REGION Network 13: Manual mode request
   RUNG wire#powerrail
      Contact( "Z256".ST_xSelectionManualMode )
      I_Contact( "Z256".ST_xManualModeAccepted )
      Coil( "Z256".ST_xManualModeRequest )
   END_RUNG
   // the same network as SCL:
   "Z256".ST_xManualModeRequest := "Z256".ST_xSelectionManualMode AND NOT "Z256".ST_xManualModeAccepted;
END_REGION

REGION Network 14: Manual mode accepted
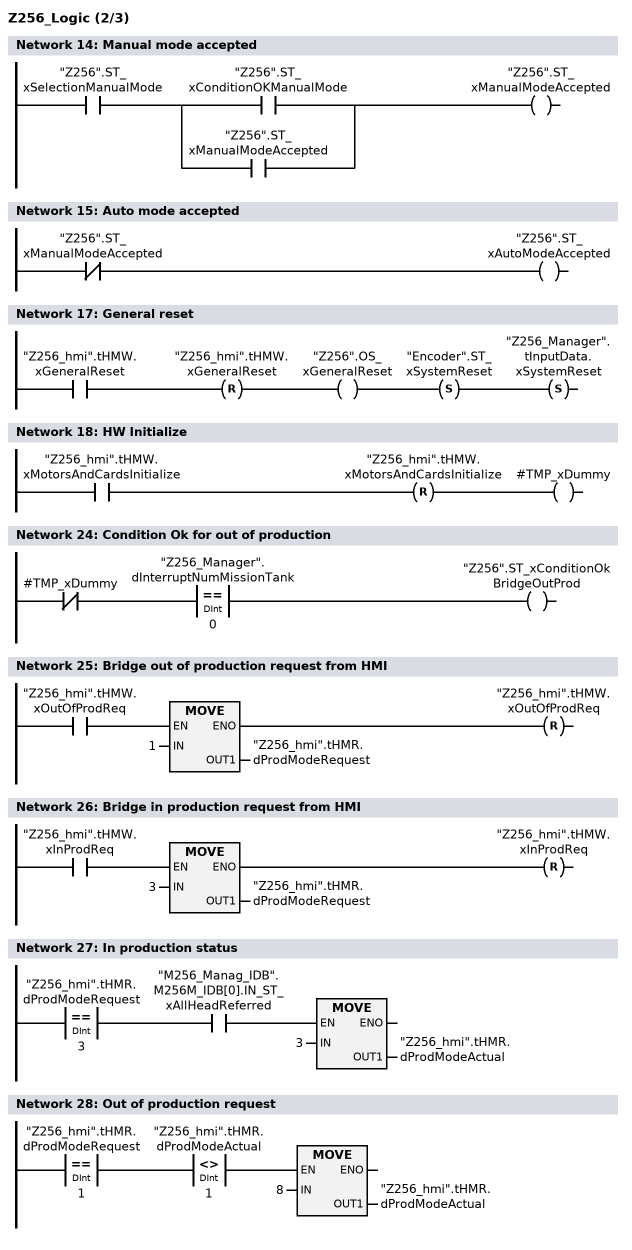
   RUNG wire#powerrail
      Contact( "Z256".ST_xSelectionManualMode )
      wire#w1
      Contact( "Z256".ST_xConditionOKManualMode )
      wire#w2
      Coil( "Z256".ST_xManualModeAccepted )
   END_RUNG
   RUNG wire#w1
      Contact( "Z256".ST_xManualModeAccepted )
   END_RUNG wire#w2
   // the same network as SCL:
   "Z256".ST_xManualModeAccepted := "Z256".ST_xSelectionManualMode AND ("Z256".ST_xConditionOKManualMode OR "Z256".ST_xManualModeAccepted);
END_REGION

REGION Network 15: Auto mode accepted
   RUNG wire#powerrail
      I_Contact( "Z256".ST_xManualModeAccepted )
      Coil( "Z256".ST_xAutoModeAccepted )
   END_RUNG
   // the same network as SCL:
   "Z256".ST_xAutoModeAccepted := NOT "Z256".ST_xManualModeAccepted;
END_REGION

REGION Network 16: ### HMI LOGICS ###
END_REGION

REGION Network 17: General reset
   RUNG wire#powerrail
      Contact( "Z256_hmi".tHMW.xGeneralReset )
      R_Coil( "Z256_hmi".tHMW.xGeneralReset )
      Coil( "Z256".OS_xGeneralReset )
      S_Coil( "Encoder".ST_xSystemReset )
      S_Coil( "Z256_Manager".tInputData.xSystemReset )
   END_RUNG
   // the same network as SCL:
   #_w1 := "Z256_hmi".tHMW.xGeneralReset;
   IF #_w1 THEN "Z256_hmi".tHMW.xGeneralReset := FALSE; END_IF;
   "Z256".OS_xGeneralReset := #_w1;
   IF #_w1 THEN
       "Encoder".ST_xSystemReset := TRUE;
       "Z256_Manager".tInputData.xSystemReset := TRUE;
   END_IF;
END_REGION

REGION Network 18: HW Initialize
   RUNG wire#powerrail
      Contact( "Z256_hmi".tHMW.xMotorsAndCardsInitialize )
      R_Coil( "Z256_hmi".tHMW.xMotorsAndCardsInitialize )
      Coil( #TMP_xDummy )
   END_RUNG
   // the same network as SCL:
   #_w1 := "Z256_hmi".tHMW.xMotorsAndCardsInitialize;
   IF #_w1 THEN "Z256_hmi".tHMW.xMotorsAndCardsInitialize := FALSE; END_IF;
   #TMP_xDummy := #_w1;
END_REGION

REGION Network 19 (SCL): Reset head initialized
   IF #TMP_xDummy THEN

       FOR #TMP_iIndex := 0 TO "CONST_dNumberOfHeadsCycle" BY 1
       DO
           "M256_Manag_IDB".M256M_IDB[#TMP_iIndex].ST_xHeadInitialized := 0;
       END_FOR;

   END_IF;
END_REGION

REGION Network 20: Cut with glass break
   // tolto enable /disable , messo che scada lo mette ad ON/OFF
END_REGION

REGION Network 21 (SCL): Enable/disable head from scada
    //   FOR #TMP_iIndex := 0 TO "CONST_dNumberOfHeadsCycle" DO
    //       IF "Z256_hmi".tHMW.rgxEnableHead[#TMP_iIndex] THEN
     //          "Z256_hmi".tHMW.rgxEnableHead[#TMP_iIndex] := 0;
     //          "Z256_hmi".tHMR.rgxHeadEnabled[#TMP_iIndex] := 1;
    //       END_IF;
    //       IF "Z256_hmi".tHMW.rgxDisableHead[#TMP_iIndex] THEN
    //           "Z256_hmi".tHMW.rgxDisableHead[#TMP_iIndex] := 0;
    //           "Z256_hmi".tHMR.rgxHeadEnabled[#TMP_iIndex] := 0;
    //       END_IF;
    //   END_FOR;
END_REGION

REGION Network 22: ### PRODUCTIONS STATUS ###
END_REGION

REGION Network 23 (SCL)
   #TMP_xDummy := false;
   FOR #TMP_iIndex:=0 TO "CONST_dNumberOfHeadsCycle" DO
       IF "Z256_Manager".tOutputData.rgxDataToProcessInter[#TMP_iIndex]=TRUE THEN
           #TMP_xDummy := true;
       END_IF;
   END_FOR;
END_REGION

REGION Network 24: Condition Ok for out of production
   RUNG wire#powerrail
      I_Contact( #TMP_xDummy )
      { S7_Templates := "SrcType := DInt" } EQ_Contact(in1 := "Z256_Manager".dInterruptNumMissionTank, in2 := 0)
      Coil( "Z256".ST_xConditionOkBridgeOutProd )
   END_RUNG
   // the same network as SCL:
   "Z256".ST_xConditionOkBridgeOutProd := NOT #TMP_xDummy AND ("Z256_Manager".dInterruptNumMissionTank = 0);
END_REGION

REGION Network 25: Bridge out of production request from HMI
   RUNG wire#powerrail
      Contact( "Z256_hmi".tHMW.xOutOfProdReq )
      Move(in := 1, out1 => "Z256_hmi".tHMR.dProdModeRequest)
      R_Coil( "Z256_hmi".tHMW.xOutOfProdReq )
   END_RUNG
   // the same network as SCL:
   IF "Z256_hmi".tHMW.xOutOfProdReq THEN
       "Z256_hmi".tHMR.dProdModeRequest := 1;
       "Z256_hmi".tHMW.xOutOfProdReq := FALSE;
   END_IF;
END_REGION

REGION Network 26: Bridge in production request from HMI
   RUNG wire#powerrail
      Contact( "Z256_hmi".tHMW.xInProdReq )
      Move(in := 3, out1 => "Z256_hmi".tHMR.dProdModeRequest)
      R_Coil( "Z256_hmi".tHMW.xInProdReq )
   END_RUNG
   // the same network as SCL:
   IF "Z256_hmi".tHMW.xInProdReq THEN
       "Z256_hmi".tHMR.dProdModeRequest := 3;
       "Z256_hmi".tHMW.xInProdReq := FALSE;
   END_IF;
END_REGION

REGION Network 27: In production status
   RUNG wire#powerrail
      { S7_Templates := "SrcType := DInt" } EQ_Contact(in1 := "Z256_hmi".tHMR.dProdModeRequest, in2 := 3)
      Contact( "M256_Manag_IDB".M256M_IDB[0].IN_ST_xAllHeadReferred )
      Move(in := 3, out1 => "Z256_hmi".tHMR.dProdModeActual)
   END_RUNG
   // the same network as SCL:
   IF ("Z256_hmi".tHMR.dProdModeRequest = 3) AND "M256_Manag_IDB".M256M_IDB[0].IN_ST_xAllHeadReferred THEN
       "Z256_hmi".tHMR.dProdModeActual := 3;
   END_IF;
END_REGION

REGION Network 28: Out of production request
   RUNG wire#powerrail
      { S7_Templates := "SrcType := DInt" } EQ_Contact(in1 := "Z256_hmi".tHMR.dProdModeRequest, in2 := 1)
      { S7_Templates := "SrcType := DInt" } NE_Contact(in1 := "Z256_hmi".tHMR.dProdModeActual, in2 := 1)
      Move(in := 8, out1 => "Z256_hmi".tHMR.dProdModeActual)
   END_RUNG
   // the same network as SCL:
   IF ("Z256_hmi".tHMR.dProdModeRequest = 1) AND ("Z256_hmi".tHMR.dProdModeActual <> 1) THEN
       "Z256_hmi".tHMR.dProdModeActual := 8;
   END_IF;
END_REGION

REGION Network 29: Out of production status
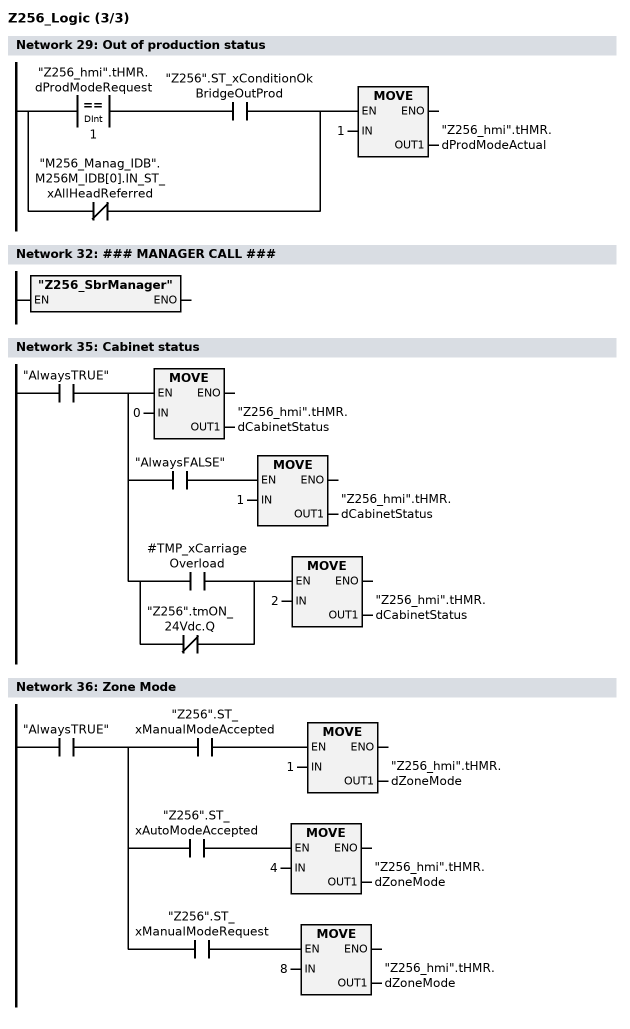
   RUNG wire#powerrail
      { S7_Templates := "SrcType := DInt" } EQ_Contact(in1 := "Z256_hmi".tHMR.dProdModeRequest, in2 := 1)
      Contact( "Z256".ST_xConditionOkBridgeOutProd )
      wire#w1
      Move(in := 1, out1 => "Z256_hmi".tHMR.dProdModeActual)
   END_RUNG
   RUNG wire#powerrail
      I_Contact( "M256_Manag_IDB".M256M_IDB[0].IN_ST_xAllHeadReferred )
   END_RUNG wire#w1
   // the same network as SCL:
   IF (("Z256_hmi".tHMR.dProdModeRequest = 1) AND "Z256".ST_xConditionOkBridgeOutProd) OR NOT "M256_Manag_IDB".M256M_IDB[0].IN_ST_xAllHeadReferred THEN
       "Z256_hmi".tHMR.dProdModeActual := 1;
   END_IF;
END_REGION

REGION Network 30 (SCL): Calculate head status

   FOR #TMP_iIndex := 0 TO "CONST_dNumberOfHeadsCycle" BY 1
   DO
       "Z256_SbrHeadsStatuses"(#TMP_iIndex);
   END_FOR;
END_REGION

REGION Network 31 (SCL): Reset head referred after emergency
   FOR #TMP_iIndex := 0 TO "CONST_dNumberOfHeadsCycle" DO
       IF "DB_Z256_Scada".tAlm.tE.x0 OR "DB_Z256_Scada".tAlm.tE.x1 OR NOT("M256_Manag_IDB".M256M_IDB[#TMP_iIndex].INPUT_xCarriageOverload) THEN
           "M256_Manag_IDB".M256M_IDB[#TMP_iIndex].ST_xHeadReferredSwitch := 0;
       END_IF;
   END_FOR;
END_REGION

REGION Network 32: ### MANAGER CALL ###
   RUNG wire#powerrail
      "Z256_SbrManager"()
   END_RUNG
   // the same network as SCL:
   "Z256_SbrManager"();
END_REGION

REGION Network 33: #### HMI STATUS ####
END_REGION

REGION Network 34 (SCL): Carriage overload array check
   #TMP_xCarriageOverload := false;
   FOR #TMP_iIndex := 0 TO "CONST_dNumberOfHeadsCycle" DO
       IF "M256_Manag_IDB".M256M_IDB[#TMP_iIndex].tALM.tS.x3 THEN
           #TMP_xCarriageOverload := true;
       END_IF;
   END_FOR;
END_REGION

REGION Network 35: Cabinet status
   RUNG wire#powerrail
      Contact( "AlwaysTRUE" )
      wire#w1
      Move(in := 0, out1 => "Z256_hmi".tHMR.dCabinetStatus)
   END_RUNG
   RUNG wire#w1
      Contact( "AlwaysFALSE" )
      Move(in := 1, out1 => "Z256_hmi".tHMR.dCabinetStatus)
   END_RUNG
   RUNG wire#w1
      Contact( #TMP_xCarriageOverload )
      wire#w2
      Move(in := 2, out1 => "Z256_hmi".tHMR.dCabinetStatus)
   END_RUNG
   RUNG wire#w1
      I_Contact( "Z256".tmON_24Vdc.Q )
   END_RUNG wire#w2
   // the same network as SCL:
   IF "AlwaysTRUE" THEN "Z256_hmi".tHMR.dCabinetStatus := 0; END_IF;
   IF "AlwaysTRUE" AND "AlwaysFALSE" THEN "Z256_hmi".tHMR.dCabinetStatus := 1; END_IF;
   IF "AlwaysTRUE" AND (#TMP_xCarriageOverload OR NOT "Z256".tmON_24Vdc.Q) THEN
       "Z256_hmi".tHMR.dCabinetStatus := 2;
   END_IF;
END_REGION

REGION Network 36: Zone Mode
   RUNG wire#powerrail
      Contact( "AlwaysTRUE" )
      wire#w1
      Contact( "Z256".ST_xManualModeAccepted )
      Move(in := 1, out1 => "Z256_hmi".tHMR.dZoneMode)
   END_RUNG
   RUNG wire#w1
      Contact( "Z256".ST_xAutoModeAccepted )
      Move(in := 4, out1 => "Z256_hmi".tHMR.dZoneMode)
   END_RUNG
   RUNG wire#w1
      Contact( "Z256".ST_xManualModeRequest )
      Move(in := 8, out1 => "Z256_hmi".tHMR.dZoneMode)
   END_RUNG
   // the same network as SCL:
   IF "AlwaysTRUE" AND "Z256".ST_xManualModeAccepted THEN "Z256_hmi".tHMR.dZoneMode := 1; END_IF;
   IF "AlwaysTRUE" AND "Z256".ST_xAutoModeAccepted THEN "Z256_hmi".tHMR.dZoneMode := 4; END_IF;
   IF "AlwaysTRUE" AND "Z256".ST_xManualModeRequest THEN "Z256_hmi".tHMR.dZoneMode := 8; END_IF;
END_REGION

REGION Network 37 (SCL): Set all brake engage/release
   IF "Z256_hmi".tHMW.tManCmd.xBrakeEngage THEN
       FOR #TMP_iIndex := 0 TO "CONST_dNumberOfHeadsCycle" BY 1
       DO
           "M256_Manag_IDB".M256M_IDB[#TMP_iIndex].tHMW.xBrakeEngageHeads := 1;
       END_FOR;
       "Z256_hmi".tHMW.tManCmd.xBrakeEngage := 0;
   END_IF;
   IF "Z256_hmi".tHMW.tManCmd.xBrakeRelease THEN
       FOR #TMP_iIndex := 0 TO "CONST_dNumberOfHeadsCycle" BY 1
       DO
           "M256_Manag_IDB".M256M_IDB[#TMP_iIndex].tHMW.xBrakeRealeaseHeads := 1;
       END_FOR;
       "Z256_hmi".tHMW.tManCmd.xBrakeRelease := 0;
   END_IF;
END_REGION
END_FUNCTION

FUNCTION "Z256_Faults" : Void   // FC3, LAD
{ S7_Optimized_Access := 'TRUE' }
VERSION : 0.1
   VAR_TEMP
      TMP_dIndex : DInt;
      TMP_dwDummy : DWord;
      TMP_dwDummy_1 : DWord;
      TMP_dwDummy_2 : DWord;
      TMP_dwDummy_3 : DWord;
      TMP_idummy : Int;
   END_VAR
   VAR_TEMP   // added for the SCL form of the ladder/FBD networks
      _w1 : Bool;
   END_VAR
BEGIN

REGION Network 1: ##### FAULTS #####
END_REGION

REGION Network 2: Reset faults
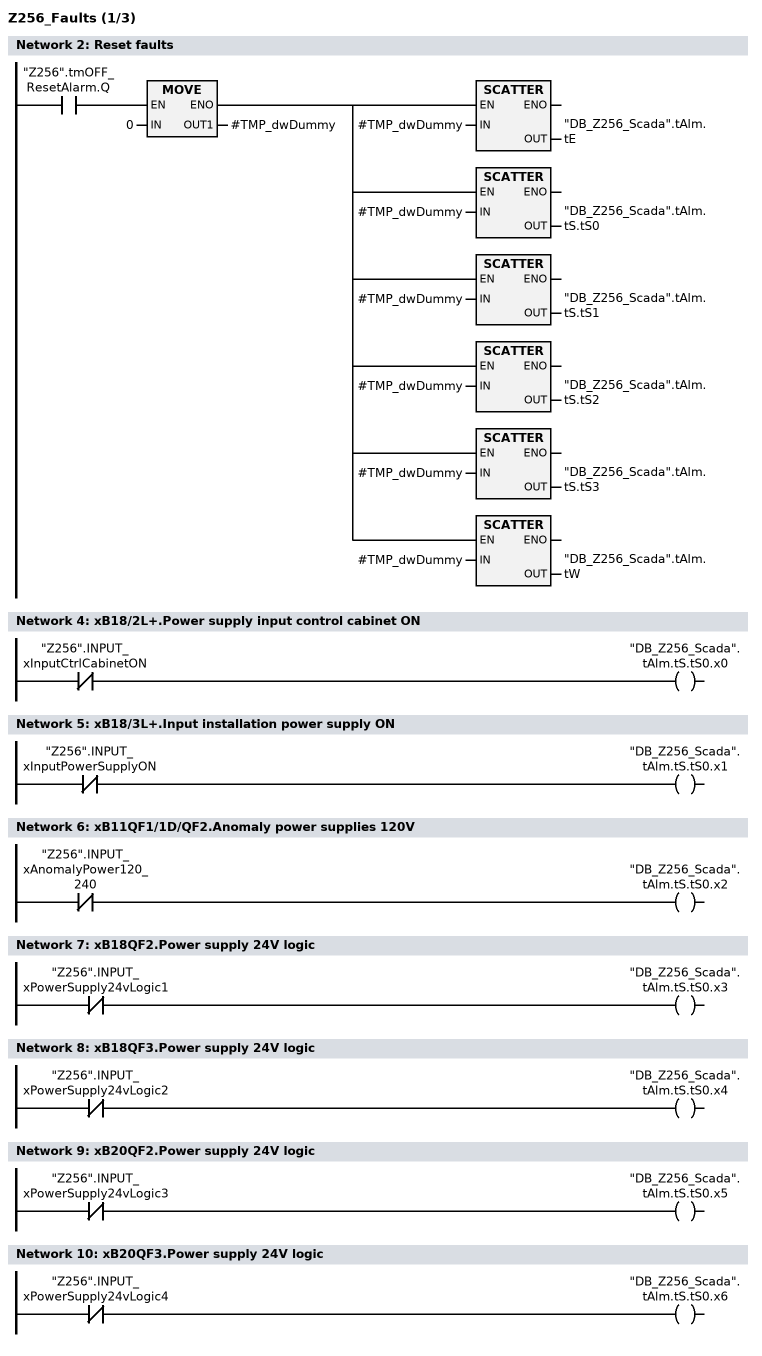
   IF "Z256".tmOFF_ResetAlarm.Q THEN #TMP_dwDummy := 0; END_IF;
   #_w1 := "Z256".tmOFF_ResetAlarm.Q;
   IF #_w1 THEN
       SCATTER(IN := #TMP_dwDummy, OUT => "DB_Z256_Scada".tAlm.tE);
       SCATTER(IN := #TMP_dwDummy, OUT => "DB_Z256_Scada".tAlm.tS.tS0);
       SCATTER(IN := #TMP_dwDummy, OUT => "DB_Z256_Scada".tAlm.tS.tS1);
       SCATTER(IN := #TMP_dwDummy, OUT => "DB_Z256_Scada".tAlm.tS.tS2);
       SCATTER(IN := #TMP_dwDummy, OUT => "DB_Z256_Scada".tAlm.tS.tS3);
       SCATTER(IN := #TMP_dwDummy, OUT => "DB_Z256_Scada".tAlm.tW);
   END_IF;
END_REGION

REGION Network 3: ### CABINET POWER FAULTS ###
END_REGION

REGION Network 4: xB18/2L+.Power supply input control cabinet ON
   RUNG wire#powerrail
      I_Contact( "Z256".INPUT_xInputCtrlCabinetON )
      Coil( "DB_Z256_Scada".tAlm.tS.tS0.x0 )
   END_RUNG
   // the same network as SCL:
   "DB_Z256_Scada".tAlm.tS.tS0.x0 := NOT "Z256".INPUT_xInputCtrlCabinetON;
END_REGION

REGION Network 5: xB18/3L+.Input installation power supply ON
   RUNG wire#powerrail
      I_Contact( "Z256".INPUT_xInputPowerSupplyON )
      Coil( "DB_Z256_Scada".tAlm.tS.tS0.x1 )
   END_RUNG
   // the same network as SCL:
   "DB_Z256_Scada".tAlm.tS.tS0.x1 := NOT "Z256".INPUT_xInputPowerSupplyON;
END_REGION

REGION Network 6: xB11QF1/1D/QF2.Anomaly power supplies 120V
   RUNG wire#powerrail
      I_Contact( "Z256".INPUT_xAnomalyPower120_240 )
      Coil( "DB_Z256_Scada".tAlm.tS.tS0.x2 )
   END_RUNG
   // the same network as SCL:
   "DB_Z256_Scada".tAlm.tS.tS0.x2 := NOT "Z256".INPUT_xAnomalyPower120_240;
END_REGION

REGION Network 7: xB18QF2.Power supply 24V logic
   RUNG wire#powerrail
      I_Contact( "Z256".INPUT_xPowerSupply24vLogic1 )
      Coil( "DB_Z256_Scada".tAlm.tS.tS0.x3 )
   END_RUNG
   // the same network as SCL:
   "DB_Z256_Scada".tAlm.tS.tS0.x3 := NOT "Z256".INPUT_xPowerSupply24vLogic1;
END_REGION

REGION Network 8: xB18QF3.Power supply 24V logic
   RUNG wire#powerrail
      I_Contact( "Z256".INPUT_xPowerSupply24vLogic2 )
      Coil( "DB_Z256_Scada".tAlm.tS.tS0.x4 )
   END_RUNG
   // the same network as SCL:
   "DB_Z256_Scada".tAlm.tS.tS0.x4 := NOT "Z256".INPUT_xPowerSupply24vLogic2;
END_REGION

REGION Network 9: xB20QF2.Power supply 24V logic
   RUNG wire#powerrail
      I_Contact( "Z256".INPUT_xPowerSupply24vLogic3 )
      Coil( "DB_Z256_Scada".tAlm.tS.tS0.x5 )
   END_RUNG
   // the same network as SCL:
   "DB_Z256_Scada".tAlm.tS.tS0.x5 := NOT "Z256".INPUT_xPowerSupply24vLogic3;
END_REGION

REGION Network 10: xB20QF3.Power supply 24V logic
   RUNG wire#powerrail
      I_Contact( "Z256".INPUT_xPowerSupply24vLogic4 )
      Coil( "DB_Z256_Scada".tAlm.tS.tS0.x6 )
   END_RUNG
   // the same network as SCL:
   "DB_Z256_Scada".tAlm.tS.tS0.x6 := NOT "Z256".INPUT_xPowerSupply24vLogic4;
END_REGION

REGION Network 11: xB21QF1.Power supply 24V logic
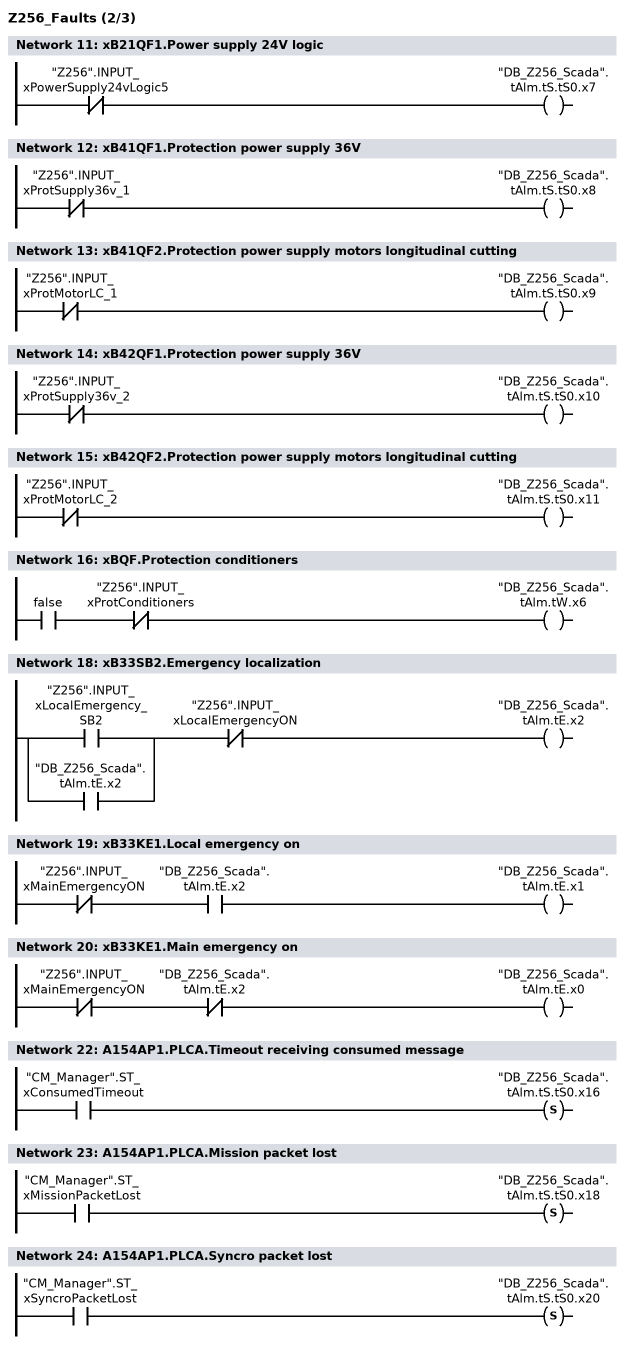
   RUNG wire#powerrail
      I_Contact( "Z256".INPUT_xPowerSupply24vLogic5 )
      Coil( "DB_Z256_Scada".tAlm.tS.tS0.x7 )
   END_RUNG
   // the same network as SCL:
   "DB_Z256_Scada".tAlm.tS.tS0.x7 := NOT "Z256".INPUT_xPowerSupply24vLogic5;
END_REGION

REGION Network 12: xB41QF1.Protection power supply 36V
   RUNG wire#powerrail
      I_Contact( "Z256".INPUT_xProtSupply36v_1 )
      Coil( "DB_Z256_Scada".tAlm.tS.tS0.x8 )
   END_RUNG
   // the same network as SCL:
   "DB_Z256_Scada".tAlm.tS.tS0.x8 := NOT "Z256".INPUT_xProtSupply36v_1;
END_REGION

REGION Network 13: xB41QF2.Protection power supply motors longitudinal cutting
   RUNG wire#powerrail
      I_Contact( "Z256".INPUT_xProtMotorLC_1 )
      Coil( "DB_Z256_Scada".tAlm.tS.tS0.x9 )
   END_RUNG
   // the same network as SCL:
   "DB_Z256_Scada".tAlm.tS.tS0.x9 := NOT "Z256".INPUT_xProtMotorLC_1;
END_REGION

REGION Network 14: xB42QF1.Protection power supply 36V
   RUNG wire#powerrail
      I_Contact( "Z256".INPUT_xProtSupply36v_2 )
      Coil( "DB_Z256_Scada".tAlm.tS.tS0.x10 )
   END_RUNG
   // the same network as SCL:
   "DB_Z256_Scada".tAlm.tS.tS0.x10 := NOT "Z256".INPUT_xProtSupply36v_2;
END_REGION

REGION Network 15: xB42QF2.Protection power supply motors longitudinal cutting
   RUNG wire#powerrail
      I_Contact( "Z256".INPUT_xProtMotorLC_2 )
      Coil( "DB_Z256_Scada".tAlm.tS.tS0.x11 )
   END_RUNG
   // the same network as SCL:
   "DB_Z256_Scada".tAlm.tS.tS0.x11 := NOT "Z256".INPUT_xProtMotorLC_2;
END_REGION

REGION Network 16: xBQF.Protection conditioners
   RUNG wire#powerrail
      Contact( false )
      I_Contact( "Z256".INPUT_xProtConditioners )
      Coil( "DB_Z256_Scada".tAlm.tW.x6 )
   END_RUNG
   // the same network as SCL:
   "DB_Z256_Scada".tAlm.tW.x6 := false AND NOT "Z256".INPUT_xProtConditioners;
END_REGION

REGION Network 17: ### EMERGENCY ###
END_REGION

REGION Network 18: xB33SB2.Emergency localization
   RUNG wire#powerrail
      Contact( "Z256".INPUT_xLocalEmergency_SB2 )
      wire#w1
      I_Contact( "Z256".INPUT_xLocalEmergencyON )
      Coil( "DB_Z256_Scada".tAlm.tE.x2 )
   END_RUNG
   RUNG wire#powerrail
      Contact( "DB_Z256_Scada".tAlm.tE.x2 )
   END_RUNG wire#w1
   // the same network as SCL:
   "DB_Z256_Scada".tAlm.tE.x2 := ("Z256".INPUT_xLocalEmergency_SB2 OR "DB_Z256_Scada".tAlm.tE.x2) AND NOT "Z256".INPUT_xLocalEmergencyON;
END_REGION

REGION Network 19: xB33KE1.Local emergency on
   RUNG wire#powerrail
      I_Contact( "Z256".INPUT_xMainEmergencyON )
      Contact( "DB_Z256_Scada".tAlm.tE.x2 )
      Coil( "DB_Z256_Scada".tAlm.tE.x1 )
   END_RUNG
   // the same network as SCL:
   "DB_Z256_Scada".tAlm.tE.x1 := NOT "Z256".INPUT_xMainEmergencyON AND "DB_Z256_Scada".tAlm.tE.x2;
END_REGION

REGION Network 20: xB33KE1.Main emergency on
   RUNG wire#powerrail
      I_Contact( "Z256".INPUT_xMainEmergencyON )
      I_Contact( "DB_Z256_Scada".tAlm.tE.x2 )
      Coil( "DB_Z256_Scada".tAlm.tE.x0 )
   END_RUNG
   // the same network as SCL:
   "DB_Z256_Scada".tAlm.tE.x0 := NOT "Z256".INPUT_xMainEmergencyON AND NOT "DB_Z256_Scada".tAlm.tE.x2;
END_REGION

REGION Network 21: ### COMMUNICATIONS STOPPING ###
END_REGION

REGION Network 22: A154AP1.PLCA.Timeout receiving consumed message
   RUNG wire#powerrail
      Contact( "CM_Manager".ST_xConsumedTimeout )
      S_Coil( "DB_Z256_Scada".tAlm.tS.tS0.x16 )
   END_RUNG
   // the same network as SCL:
   IF "CM_Manager".ST_xConsumedTimeout THEN "DB_Z256_Scada".tAlm.tS.tS0.x16 := TRUE; END_IF;
END_REGION

REGION Network 23: A154AP1.PLCA.Mission packet lost
   RUNG wire#powerrail
      Contact( "CM_Manager".ST_xMissionPacketLost )
      S_Coil( "DB_Z256_Scada".tAlm.tS.tS0.x18 )
   END_RUNG
   // the same network as SCL:
   IF "CM_Manager".ST_xMissionPacketLost THEN "DB_Z256_Scada".tAlm.tS.tS0.x18 := TRUE; END_IF;
END_REGION

REGION Network 24: A154AP1.PLCA.Syncro packet lost
   RUNG wire#powerrail
      Contact( "CM_Manager".ST_xSyncroPacketLost )
      S_Coil( "DB_Z256_Scada".tAlm.tS.tS0.x20 )
   END_RUNG
   // the same network as SCL:
   IF "CM_Manager".ST_xSyncroPacketLost THEN "DB_Z256_Scada".tAlm.tS.tS0.x20 := TRUE; END_IF;
END_REGION

REGION Network 25: ### SYNCRONIZATION ###
END_REGION

REGION Network 26: Syncro.YCut meter gap outside the limits
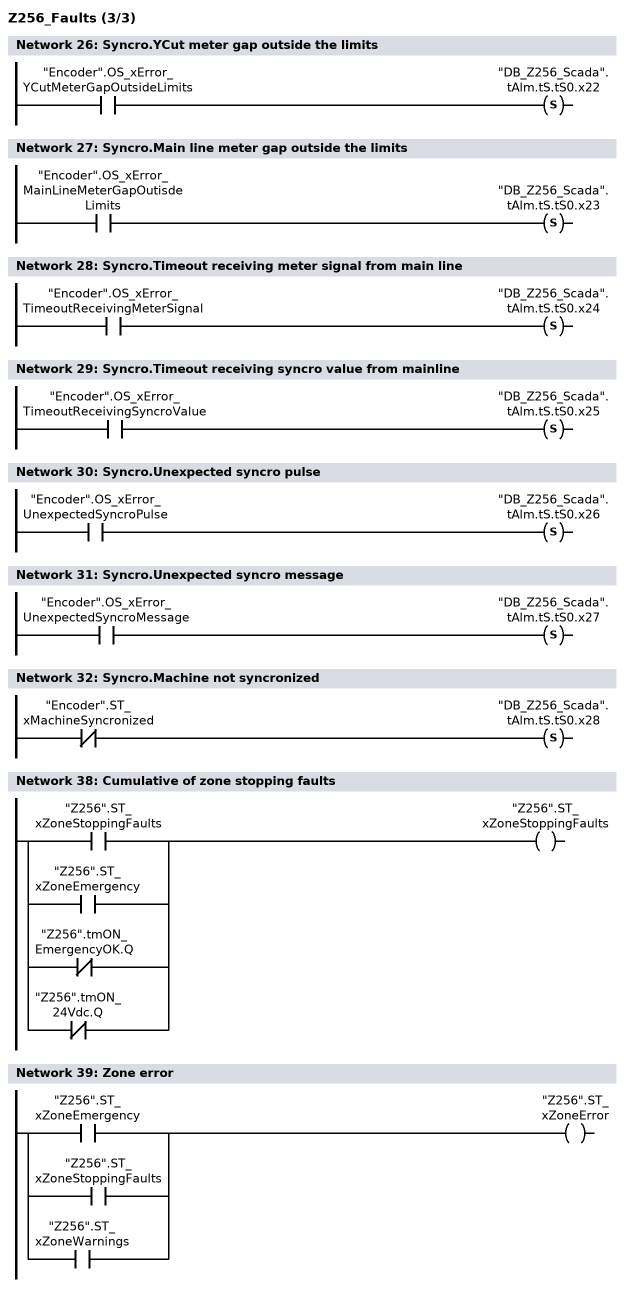
   RUNG wire#powerrail
      Contact( "Encoder".OS_xError_YCutMeterGapOutsideLimits )
      S_Coil( "DB_Z256_Scada".tAlm.tS.tS0.x22 )
   END_RUNG
   // the same network as SCL:
   IF "Encoder".OS_xError_YCutMeterGapOutsideLimits THEN "DB_Z256_Scada".tAlm.tS.tS0.x22 := TRUE; END_IF;
END_REGION

REGION Network 27: Syncro.Main line meter gap outside the limits
   RUNG wire#powerrail
      Contact( "Encoder".OS_xError_MainLineMeterGapOutisdeLimits )
      S_Coil( "DB_Z256_Scada".tAlm.tS.tS0.x23 )
   END_RUNG
   // the same network as SCL:
   IF "Encoder".OS_xError_MainLineMeterGapOutisdeLimits THEN "DB_Z256_Scada".tAlm.tS.tS0.x23 := TRUE; END_IF;
END_REGION

REGION Network 28: Syncro.Timeout receiving meter signal from main line
   RUNG wire#powerrail
      Contact( "Encoder".OS_xError_TimeoutReceivingMeterSignal )
      S_Coil( "DB_Z256_Scada".tAlm.tS.tS0.x24 )
   END_RUNG
   // the same network as SCL:
   IF "Encoder".OS_xError_TimeoutReceivingMeterSignal THEN "DB_Z256_Scada".tAlm.tS.tS0.x24 := TRUE; END_IF;
END_REGION

REGION Network 29: Syncro.Timeout receiving syncro value from mainline
   RUNG wire#powerrail
      Contact( "Encoder".OS_xError_TimeoutReceivingSyncroValue )
      S_Coil( "DB_Z256_Scada".tAlm.tS.tS0.x25 )
   END_RUNG
   // the same network as SCL:
   IF "Encoder".OS_xError_TimeoutReceivingSyncroValue THEN "DB_Z256_Scada".tAlm.tS.tS0.x25 := TRUE; END_IF;
END_REGION

REGION Network 30: Syncro.Unexpected syncro pulse
   RUNG wire#powerrail
      Contact( "Encoder".OS_xError_UnexpectedSyncroPulse )
      S_Coil( "DB_Z256_Scada".tAlm.tS.tS0.x26 )
   END_RUNG
   // the same network as SCL:
   IF "Encoder".OS_xError_UnexpectedSyncroPulse THEN "DB_Z256_Scada".tAlm.tS.tS0.x26 := TRUE; END_IF;
END_REGION

REGION Network 31: Syncro.Unexpected syncro message
   RUNG wire#powerrail
      Contact( "Encoder".OS_xError_UnexpectedSyncroMessage )
      S_Coil( "DB_Z256_Scada".tAlm.tS.tS0.x27 )
   END_RUNG
   // the same network as SCL:
   IF "Encoder".OS_xError_UnexpectedSyncroMessage THEN "DB_Z256_Scada".tAlm.tS.tS0.x27 := TRUE; END_IF;
END_REGION

REGION Network 32: Syncro.Machine not syncronized
   RUNG wire#powerrail
      I_Contact( "Encoder".ST_xMachineSyncronized )
      S_Coil( "DB_Z256_Scada".tAlm.tS.tS0.x28 )
   END_RUNG
   // the same network as SCL:
   IF NOT "Encoder".ST_xMachineSyncronized THEN "DB_Z256_Scada".tAlm.tS.tS0.x28 := TRUE; END_IF;
END_REGION

REGION Network 33: ### CUMULATIVE BITS ###
END_REGION

REGION Network 34 (SCL): Cumulative of emergency faults active
   "Z256".ST_xZoneEmergency := 0;

   GATHER(IN:= "DB_Z256_Scada".tAlm.tE,
          OUT=>#TMP_dwDummy);

   IF #TMP_dwDummy <> 0 THEN
       "Z256".ST_xZoneEmergency := 1;
   END_IF;
END_REGION

REGION Network 35 (SCL): Cumulative of warning active
   "Z256".ST_xZoneWarnings := 0;

   GATHER(IN:= "DB_Z256_Scada".tAlm.tW,
          OUT=>#TMP_dwDummy);

   IF #TMP_dwDummy <> 0 THEN
       "Z256".ST_xZoneWarnings := 1;
   END_IF;
END_REGION

REGION Network 36 (SCL): Cumulative of stopping faults active
   "Z256".ST_xZoneStoppingFaults := 0;
   GATHER(IN := "DB_Z256_Scada".tAlm.tS.tS0,
          OUT => #TMP_dwDummy);
   GATHER(IN := "DB_Z256_Scada".tAlm.tS.tS1,
          OUT => #TMP_dwDummy_1);
   GATHER(IN := "DB_Z256_Scada".tAlm.tS.tS2,
          OUT => #TMP_dwDummy_2);
   GATHER(IN := "DB_Z256_Scada".tAlm.tS.tS3,
          OUT => #TMP_dwDummy_3);

   IF #TMP_dwDummy <> 0 AND #TMP_dwDummy_1 <> 0 AND #TMP_dwDummy_2 <> 0 AND #TMP_dwDummy_3 <> 0  THEN
       "Z256".ST_xZoneStoppingFaults := 1;
   END_IF;
END_REGION

REGION Network 37 (SCL): Cumulative of faults active
   "Z256".ST_xZoneFaults := 0;
   GATHER(IN := "DB_Z256_Scada".tAlm.tF,
          OUT => #TMP_dwDummy);

   IF #TMP_dwDummy <> 0 THEN
       "Z256".ST_xZoneFaults := 1;
   END_IF;
END_REGION

REGION Network 38: Cumulative of zone stopping faults
   RUNG wire#powerrail
      Contact( "Z256".ST_xZoneStoppingFaults )
      wire#w1
      Coil( "Z256".ST_xZoneStoppingFaults )
   END_RUNG
   RUNG wire#powerrail
      Contact( "Z256".ST_xZoneEmergency )
   END_RUNG wire#w1
   RUNG wire#powerrail
      I_Contact( "Z256".tmON_EmergencyOK.Q )
   END_RUNG wire#w1
   RUNG wire#powerrail
      I_Contact( "Z256".tmON_24Vdc.Q )
   END_RUNG wire#w1
   // the same network as SCL:
   "Z256".ST_xZoneStoppingFaults := "Z256".ST_xZoneStoppingFaults OR "Z256".ST_xZoneEmergency OR NOT "Z256".tmON_EmergencyOK.Q OR NOT "Z256".tmON_24Vdc.Q;
END_REGION

REGION Network 39: Zone error
   RUNG wire#powerrail
      Contact( "Z256".ST_xZoneEmergency )
      wire#w1
      Coil( "Z256".ST_xZoneError )
   END_RUNG
   RUNG wire#powerrail
      Contact( "Z256".ST_xZoneStoppingFaults )
   END_RUNG wire#w1
   RUNG wire#powerrail
      Contact( "Z256".ST_xZoneWarnings )
   END_RUNG wire#w1
   // the same network as SCL:
   "Z256".ST_xZoneError := "Z256".ST_xZoneEmergency OR "Z256".ST_xZoneStoppingFaults OR "Z256".ST_xZoneWarnings;
END_REGION
END_FUNCTION

FUNCTION "Z256_SbrHeadsStatuses" : Void   // FC4, LAD
{ S7_Optimized_Access := 'TRUE' }
VERSION : 0.1
   VAR_INPUT
      IN_Index : Int;
   END_VAR
BEGIN

REGION Network 1: #### CALCULATE HEAD STATUSES ####
END_REGION

REGION Network 2: Condition OK head out of service - ###TEMP###
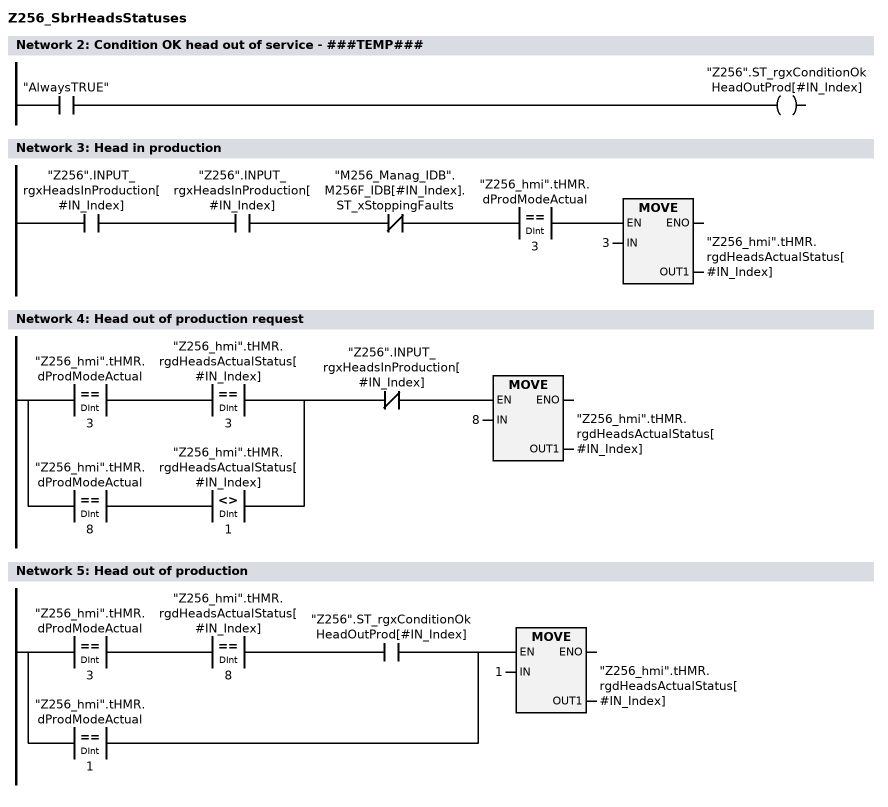
   RUNG wire#powerrail
      Contact( "AlwaysTRUE" )
      Coil( "Z256".ST_rgxConditionOkHeadOutProd[#IN_Index] )
   END_RUNG
   // the same network as SCL:
   "Z256".ST_rgxConditionOkHeadOutProd[#IN_Index] := "AlwaysTRUE";
END_REGION

REGION Network 3: Head in production
   RUNG wire#powerrail
      Contact( "Z256".INPUT_rgxHeadsInProduction[#IN_Index] )
      Contact( "Z256".INPUT_rgxHeadsInProduction[#IN_Index] )
      I_Contact( "M256_Manag_IDB".M256F_IDB[#IN_Index].ST_xStoppingFaults )
      { S7_Templates := "SrcType := DInt" } EQ_Contact(in1 := "Z256_hmi".tHMR.dProdModeActual, in2 := 3)
      Move(in := 3, out1 => "Z256_hmi".tHMR.rgdHeadsActualStatus[#IN_Index])
   END_RUNG
   // the same network as SCL:
   IF "Z256".INPUT_rgxHeadsInProduction[#IN_Index] AND "Z256".INPUT_rgxHeadsInProduction[#IN_Index] AND NOT "M256_Manag_IDB".M256F_IDB[#IN_Index].ST_xStoppingFaults AND ("Z256_hmi".tHMR.dProdModeActual = 3) THEN
       "Z256_hmi".tHMR.rgdHeadsActualStatus[#IN_Index] := 3;
   END_IF;
END_REGION

REGION Network 4: Head out of production request
   RUNG wire#powerrail
      { S7_Templates := "SrcType := DInt" } EQ_Contact(in1 := "Z256_hmi".tHMR.dProdModeActual, in2 := 3)
      { S7_Templates := "SrcType := DInt" } EQ_Contact(in1 := "Z256_hmi".tHMR.rgdHeadsActualStatus[#IN_Index], in2 := 3)
      wire#w1
      I_Contact( "Z256".INPUT_rgxHeadsInProduction[#IN_Index] )
      Move(in := 8, out1 => "Z256_hmi".tHMR.rgdHeadsActualStatus[#IN_Index])
   END_RUNG
   RUNG wire#powerrail
      { S7_Templates := "SrcType := DInt" } EQ_Contact(in1 := "Z256_hmi".tHMR.dProdModeActual, in2 := 8)
      { S7_Templates := "SrcType := DInt" } NE_Contact(in1 := "Z256_hmi".tHMR.rgdHeadsActualStatus[#IN_Index], in2 := 1)
   END_RUNG wire#w1
   // the same network as SCL:
   IF ((("Z256_hmi".tHMR.dProdModeActual = 3) AND ("Z256_hmi".tHMR.rgdHeadsActualStatus[#IN_Index] = 3)) OR (("Z256_hmi".tHMR.dProdModeActual = 8) AND ("Z256_hmi".tHMR.rgdHeadsActualStatus[#IN_Index] <> 1))) AND NOT "Z256".INPUT_rgxHeadsInProduction[#IN_Index] THEN
       "Z256_hmi".tHMR.rgdHeadsActualStatus[#IN_Index] := 8;
   END_IF;
END_REGION

REGION Network 5: Head out of production
   RUNG wire#powerrail
      { S7_Templates := "SrcType := DInt" } EQ_Contact(in1 := "Z256_hmi".tHMR.dProdModeActual, in2 := 3)
      { S7_Templates := "SrcType := DInt" } EQ_Contact(in1 := "Z256_hmi".tHMR.rgdHeadsActualStatus[#IN_Index], in2 := 8)
      Contact( "Z256".ST_rgxConditionOkHeadOutProd[#IN_Index] )
      wire#w1
      Move(in := 1, out1 => "Z256_hmi".tHMR.rgdHeadsActualStatus[#IN_Index])
   END_RUNG
   RUNG wire#powerrail
      { S7_Templates := "SrcType := DInt" } EQ_Contact(in1 := "Z256_hmi".tHMR.dProdModeActual, in2 := 1)
   END_RUNG wire#w1
   // the same network as SCL:
   IF (("Z256_hmi".tHMR.dProdModeActual = 3) AND ("Z256_hmi".tHMR.rgdHeadsActualStatus[#IN_Index] = 8) AND "Z256".ST_rgxConditionOkHeadOutProd[#IN_Index]) OR ("Z256_hmi".tHMR.dProdModeActual = 1) THEN
       "Z256_hmi".tHMR.rgdHeadsActualStatus[#IN_Index] := 1;
   END_IF;
END_REGION
END_FUNCTION

FUNCTION "Z256_SbrManager" : Void   // FC5, SCL
{ S7_Optimized_Access := 'TRUE' }
VERSION : 0.1
   VAR_TEMP
      TMP_dIndex : DInt;
      TMP_xOutputMergeMission : Bool;
      TMP_dDummy : DInt;
      TMP_dInsideIndex : DInt;
      TMP_xCheckNext : Bool;
      TMP_dLineOverlap : DInt;
      TMP_xProcNextAllowed : Bool;
      TMP_xIsDiffent : Bool;
      TMP_xDummy : Bool;
      TMP_dSize : DInt;
      TMP_dIndex2 : DInt;
      TMP_dSize2 : DInt;
      TMP_dIndex3 : DInt;
      TMP_vVariant : Variant;
      n : DInt;
      TMP_iReturn : Int;
   END_VAR
BEGIN
   ////--------------------------------------------------------------------------------------------------------------------
   //   Copyright (c)  Bottero Spa
   //--------------------------------------------------------------
   //   Routine: YCUT Manager
   //       Author: Elia Lerda
   //   Created: May-2018
   //--------------------------------------------------------------
   //   Description: This routine will manage all the mission to the YCUT bridge
   //
   //   History:
   //
   ////--------------------------------------------------------------------------------------------------------------------


   //MAPPING THE INPUT DATA TO THE PROCEDURE

   FOR #TMP_dIndex := 0 TO "CONST_dNumberOfHeadsCycle" DO

       "Z256_Manager".tInputData.rgdArmONReaction_ms[#TMP_dIndex] := "M256_Manag_IDB".M256A_IDB[#TMP_dIndex].tHMW.dDescentReactTime_ms + 200;
       "Z256_Manager".tInputData.rgdArmOFFReaction_ms[#TMP_dIndex] := "M256_Manag_IDB".M256A_IDB[#TMP_dIndex].tHMW.dRaiseReactTime_ms;
       "Z256_Manager".tInputData.rgdFireONReaction_ms[#TMP_dIndex] := "M256_Manag_IDB".M256F_IDB[#TMP_dIndex].tHMW.dHeadFireONReaction_ms;
       "Z256_Manager".tInputData.rgdFireOFFReaction_ms[#TMP_dIndex] := "M256_Manag_IDB".M256F_IDB[#TMP_dIndex].tHMW.dHeadFireOFFReaction_ms;
       "Z256_Manager".tInputData.rgdOilDelayStart_ms[#TMP_dIndex] := "M256_Manag_IDB".M256F_IDB[#TMP_dIndex].tHMW.dHeadOilONDelay_ms;
       "Z256_Manager".tInputData.rgdOilDelayEnd_ms[#TMP_dIndex] := "M256_Manag_IDB".M256F_IDB[#TMP_dIndex].tHMW.dHeadOilOFFDelay_ms;
       "Z256_Manager".tInputData.rgdFireONDelayStart_cmm[#TMP_dIndex] := "M256_Manag_IDB".M256F_IDB[#TMP_dIndex].tHMW.dHeadFireONDelay_cmm;
       "Z256_Manager".tInputData.rgdFireOFFDelayEnd_cmm[#TMP_dIndex] := "M256_Manag_IDB".M256F_IDB[#TMP_dIndex].tHMW.dHeadFireOFFDelay_cmm;

   END_FOR;

   //If buffer full reject any mission
   IF "Z256_Manager".dInterruptNumMissionTank >= 20 THEN

       "Z256_Manager".tInputData.xNewMission := 0;

   END_IF;


   // --- First step - Look if there are new mission to insert inside the tank ---
   IF "Z256_Manager".tInputData.xNewMission AND NOT "Z256_Manager".tOutputData.xGateOpen THEN

       //--- INSERT MISSION FOR INTERRUPT ---
       #TMP_dIndex := "Z256_Manager".dInterruptNumMissionTank;
       //TMP_dMergeID := Z256_Manager.tInputData.dMissionCode;
       #TMP_xOutputMergeMission := 0;

       IF "Z256_Manager".dInterruptNumMissionTank > 0 THEN

           //The mission tank has mission, check if the last one is nearest this mission
           #TMP_dDummy := "Z256_Manager".tInputData.dMissionStart_cmm - "Z256_Manager".rgtInterruptMissionTank["Z256_Manager".dInterruptNumMissionTank - 1].dMissionValue_cmm;

           IF ABS(#TMP_dDummy) <= "CONST_dFire_OnOff_MaxValue" THEN
               //The difference is less than the maximum offset. Merge the mission
               #TMP_dIndex := #TMP_dIndex - 1;
               //TMP_dMergeID := Z256_Manager.rgtInterruptMissionTank[TMP_dIndex].dMissionCode;
           END_IF;

       ELSE

           //If no mission on tank, check if the mission is nearest to one already
           //on the output. If yes create only the end.
           #TMP_dDummy := "Z256_Manager".tInputData.dMissionStart_cmm - "Z256_Manager".tOutputData.dTargetLineValue_cmm;

           IF ABS(#TMP_dDummy) <= "CONST_dFire_OnOff_MaxValue" THEN
               //The difference is less than the maximum offset. Merge the mission
               #TMP_xOutputMergeMission := 1;


           END_IF;